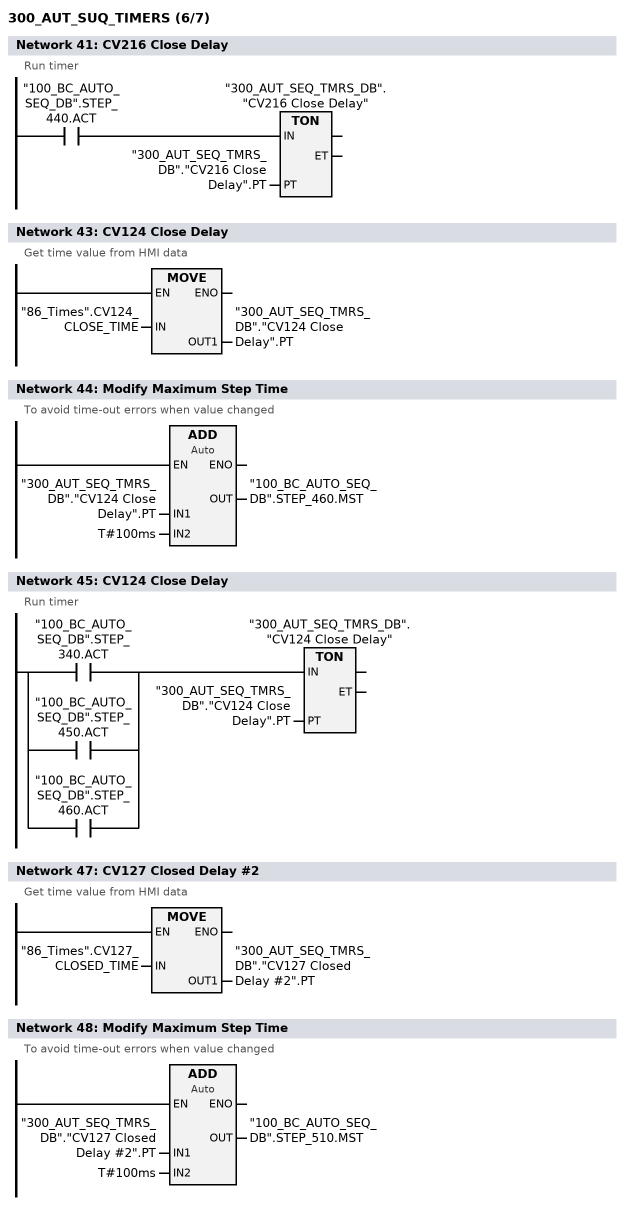
   "300_AUT_SEQ_TMRS_DB"."CV216 Close Delay".TON(IN := "100_BC_AUTO_SEQ_DB".STEP_440.ACT,
                           PT := "300_AUT_SEQ_TMRS_DB"."CV216 Close Delay".PT);
END_REGION

REGION Network 43: CV124 Close Delay
   // Get time value from HMI data
   RUNG wire#powerrail
      Move(in := "86_Times".CV124_CLOSE_TIME, out1 => "300_AUT_SEQ_TMRS_DB"."CV124 Close Delay".PT)
   END_RUNG
   // the same network as SCL:
   "300_AUT_SEQ_TMRS_DB"."CV124 Close Delay".PT := "86_Times".CV124_CLOSE_TIME;
END_REGION

REGION Network 44: Modify Maximum Step Time
   // To avoid time-out errors when value changed
   RUNG wire#powerrail
      Add(in1 := "300_AUT_SEQ_TMRS_DB"."CV124 Close Delay".PT, in2 := T#100ms, out => "100_BC_AUTO_SEQ_DB".STEP_460.MST)
   END_RUNG
   // the same network as SCL:
   "100_BC_AUTO_SEQ_DB".STEP_460.MST := "300_AUT_SEQ_TMRS_DB"."CV124 Close Delay".PT + T#100ms;
END_REGION

REGION Network 45: CV124 Close Delay
   // Run timer
   "300_AUT_SEQ_TMRS_DB"."CV124 Close Delay".TON(IN := "100_BC_AUTO_SEQ_DB".STEP_340.ACT OR "100_BC_AUTO_SEQ_DB".STEP_450.ACT OR "100_BC_AUTO_SEQ_DB".STEP_460.ACT,
                           PT := "300_AUT_SEQ_TMRS_DB"."CV124 Close Delay".PT);
END_REGION

REGION Network 47: CV127 Closed Delay #2
   // Get time value from HMI data
   RUNG wire#powerrail
      Move(in := "86_Times".CV127_CLOSED_TIME, out1 => "300_AUT_SEQ_TMRS_DB"."CV127 Closed Delay #2".PT)
   END_RUNG
   // the same network as SCL:
   "300_AUT_SEQ_TMRS_DB"."CV127 Closed Delay #2".PT := "86_Times".CV127_CLOSED_TIME;
END_REGION

REGION Network 48: Modify Maximum Step Time
   // To avoid time-out errors when value changed
   RUNG wire#powerrail
      Add(in1 := "300_AUT_SEQ_TMRS_DB"."CV127 Closed Delay #2".PT, in2 := T#100ms, out => "100_BC_AUTO_SEQ_DB".STEP_510.MST)
   END_RUNG
   // the same network as SCL:
   "100_BC_AUTO_SEQ_DB".STEP_510.MST := "300_AUT_SEQ_TMRS_DB"."CV127 Closed Delay #2".PT + T#100ms;
END_REGION

REGION Network 49: CV127 Closed Delay #2
   // Run timer
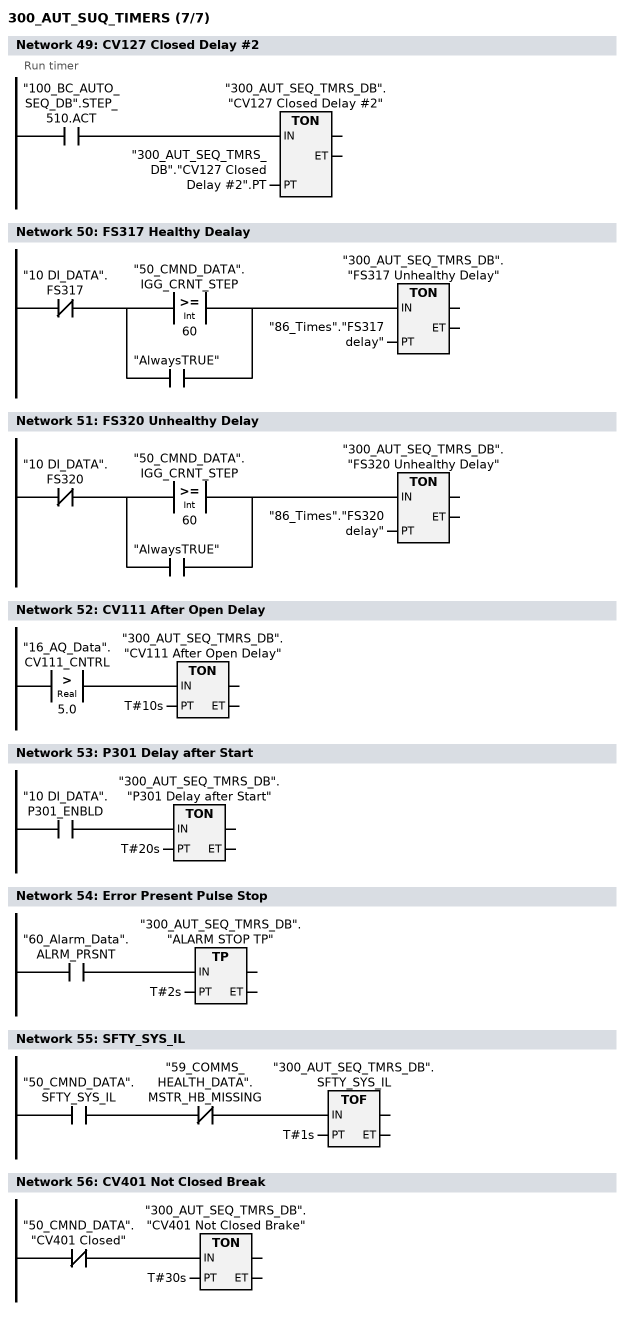
   "300_AUT_SEQ_TMRS_DB"."CV127 Closed Delay #2".TON(IN := "100_BC_AUTO_SEQ_DB".STEP_510.ACT,
                           PT := "300_AUT_SEQ_TMRS_DB"."CV127 Closed Delay #2".PT);
END_REGION

REGION Network 50: FS317 Healthy Dealay
   "300_AUT_SEQ_TMRS_DB"."FS317 Unhealthy Delay".TON(IN := NOT "10 DI_DATA".FS317 AND (("50_CMND_DATA".IGG_CRNT_STEP >= 60) OR "AlwaysTRUE"),
                           PT := "86_Times"."FS317 delay");
END_REGION

REGION Network 51: FS320 Unhealthy Delay
   "300_AUT_SEQ_TMRS_DB"."FS320 Unhealthy Delay".TON(IN := NOT "10 DI_DATA".FS320 AND (("50_CMND_DATA".IGG_CRNT_STEP >= 60) OR "AlwaysTRUE"),
                           PT := "86_Times"."FS320 delay");
END_REGION

REGION Network 52: CV111 After Open Delay
   "300_AUT_SEQ_TMRS_DB"."CV111 After Open Delay".TON(IN := "16_AQ_Data".CV111_CNTRL > 5.0, PT := T#10s);
END_REGION

REGION Network 53: P301 Delay after Start
   "300_AUT_SEQ_TMRS_DB"."P301 Delay after Start".TON(IN := "10 DI_DATA".P301_ENBLD, PT := T#20s);
END_REGION

REGION Network 54: Error Present Pulse Stop
   "300_AUT_SEQ_TMRS_DB"."ALARM STOP TP".TP(IN := "60_Alarm_Data".ALRM_PRSNT, PT := T#2s);
END_REGION

REGION Network 55: SFTY_SYS_IL
   "300_AUT_SEQ_TMRS_DB".SFTY_SYS_IL.TOF(IN := "50_CMND_DATA".SFTY_SYS_IL AND NOT "59_COMMS_HEALTH_DATA".MSTR_HB_MISSING,
                           PT := T#1s);
END_REGION

REGION Network 56: CV401 Not Closed Break
   "300_AUT_SEQ_TMRS_DB"."CV401 Not Closed Brake".TON(IN := NOT "50_CMND_DATA"."CV401 Closed", PT := T#30s);
END_REGION
END_FUNCTION

// folder: 50 - 59 PLC Communication

FUNCTION "51_GET_SLAVE_DATA" : Void   // FC51, LAD
TITLE = Get Slave Status Data
{ S7_Optimized_Access := 'TRUE' }
AUTHOR : JRS
VERSION : 0.1
// Code for getting status data from the slave PLC (IGG)
   VAR_TEMP
      RET_VAL_1 : Int;
   END_VAR
BEGIN

REGION Network 1: Get Slave Status Data
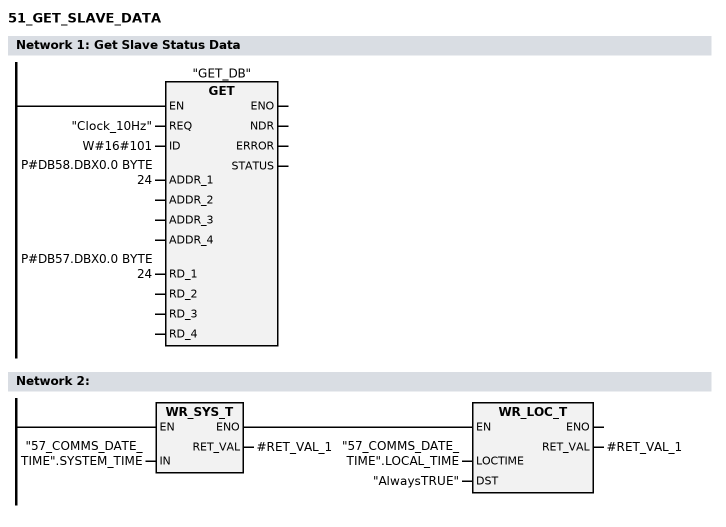
   "GET_DB"(REQ := "Clock_10Hz", ID := W#16#101, ADDR_1 := P#DB58.DBX0.0 BYTE 24, RD_1 := P#DB57.DBX0.0 BYTE 24);   // GET
END_REGION

REGION Network 2
   // ENO of a box is taken as its EN; it also drops when the box reports an error
   #RET_VAL_1 := WR_SYS_T(IN := "57_COMMS_DATE_TIME".SYSTEM_TIME);
   #RET_VAL_1 := WR_LOC_T(LOCTIME := "57_COMMS_DATE_TIME".LOCAL_TIME, DST := "AlwaysTRUE");
END_REGION
END_FUNCTION

FUNCTION "59_COMMS_HEALTH" : Void   // FC59, LAD
TITLE = Communications Heart Beats
{ S7_Optimized_Access := 'TRUE' }
AUTHOR : JRS
VERSION : 0.1
// Code for communications health determination
   VAR_TEMP   // added for the SCL form of the ladder/FBD networks
      _w1 : Bool;
   END_VAR
BEGIN

REGION Network 1: Local Heart Beat
   // Flip flop for status to other PLC's
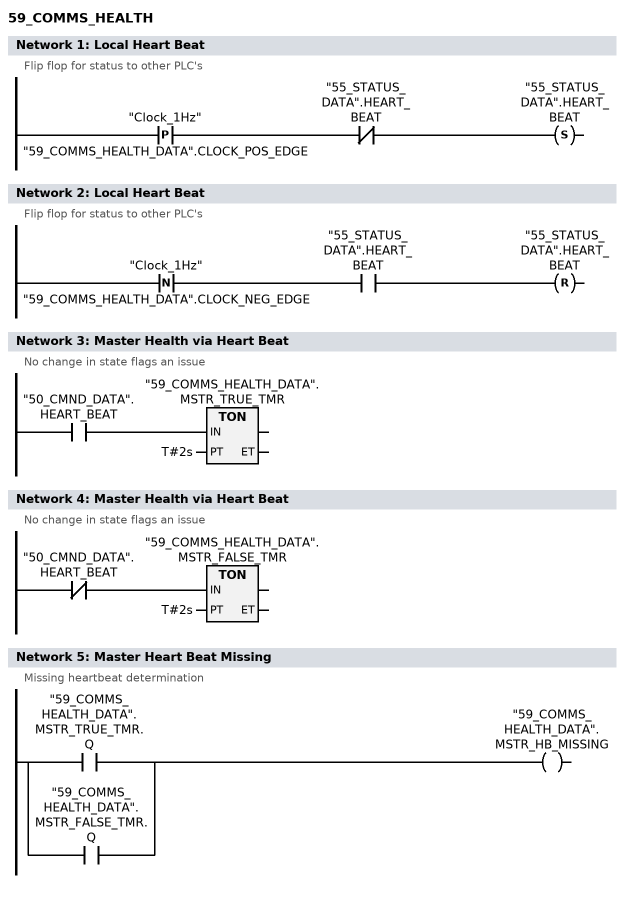
   RUNG wire#powerrail
      P_Contact(operand := "Clock_1Hz", bit := "59_COMMS_HEALTH_DATA".CLOCK_POS_EDGE)
      I_Contact( "55_STATUS_DATA".HEART_BEAT )
      S_Coil( "55_STATUS_DATA".HEART_BEAT )
   END_RUNG
   // the same network as SCL:
   #_w1 := "Clock_1Hz" AND NOT "59_COMMS_HEALTH_DATA".CLOCK_POS_EDGE;   // rising edge of "Clock_1Hz"
   "59_COMMS_HEALTH_DATA".CLOCK_POS_EDGE := "Clock_1Hz";
   IF #_w1 AND NOT "55_STATUS_DATA".HEART_BEAT THEN "55_STATUS_DATA".HEART_BEAT := TRUE; END_IF;
END_REGION

REGION Network 2: Local Heart Beat
   // Flip flop for status to other PLC's
   RUNG wire#powerrail
      N_Contact(operand := "Clock_1Hz", bit := "59_COMMS_HEALTH_DATA".CLOCK_NEG_EDGE)
      Contact( "55_STATUS_DATA".HEART_BEAT )
      R_Coil( "55_STATUS_DATA".HEART_BEAT )
   END_RUNG
   // the same network as SCL:
   #_w1 := NOT "Clock_1Hz" AND "59_COMMS_HEALTH_DATA".CLOCK_NEG_EDGE;   // falling edge of "Clock_1Hz"
   "59_COMMS_HEALTH_DATA".CLOCK_NEG_EDGE := "Clock_1Hz";
   IF #_w1 AND "55_STATUS_DATA".HEART_BEAT THEN "55_STATUS_DATA".HEART_BEAT := FALSE; END_IF;
END_REGION

REGION Network 3: Master Health via Heart Beat
   // No change in state flags an issue
   "59_COMMS_HEALTH_DATA".MSTR_TRUE_TMR.TON(IN := "50_CMND_DATA".HEART_BEAT, PT := T#2s);
END_REGION

REGION Network 4: Master Health via Heart Beat
   // No change in state flags an issue
   "59_COMMS_HEALTH_DATA".MSTR_FALSE_TMR.TON(IN := NOT "50_CMND_DATA".HEART_BEAT, PT := T#2s);
END_REGION

REGION Network 5: Master Heart Beat Missing
   // Missing heartbeat determination
   RUNG wire#powerrail
      Contact( "59_COMMS_HEALTH_DATA".MSTR_TRUE_TMR.Q )
      wire#w1
      Coil( "59_COMMS_HEALTH_DATA".MSTR_HB_MISSING )
   END_RUNG
   RUNG wire#powerrail
      Contact( "59_COMMS_HEALTH_DATA".MSTR_FALSE_TMR.Q )
   END_RUNG wire#w1
   // the same network as SCL:
   "59_COMMS_HEALTH_DATA".MSTR_HB_MISSING := "59_COMMS_HEALTH_DATA".MSTR_TRUE_TMR.Q OR "59_COMMS_HEALTH_DATA".MSTR_FALSE_TMR.Q;
END_REGION
END_FUNCTION

// folder: 500 - 699 Standard FBs

FUNCTION_BLOCK "500_SEQ_STEP"   // FB500, LAD
{ S7_Optimized_Access := 'TRUE' }
VERSION : 0.1
   VAR_INPUT
      SN : Int;   // Step number
      CS : Int;   // Current step
      MST : Time;   // Maximum step time
      SC : Bool;   // Step complete
      BPFLT : Bool;   // Bypass fault
   END_VAR
   VAR_OUTPUT
      ACT : Bool;   // Active
      DN : Bool;   // Done
   END_VAR
   VAR_IN_OUT
      AMST : Time;   // Actual maximum step time
      FLT : Bool;   // Timed out
   END_VAR
   VAR
      RNG : Bool;   // Running
   END_VAR
   VAR RETAIN
      STP_MAX_TIM : TON_TIME;   // Maximum step time
   END_VAR
BEGIN

REGION Network 1: Step Active
   // When step number is active, it is also running
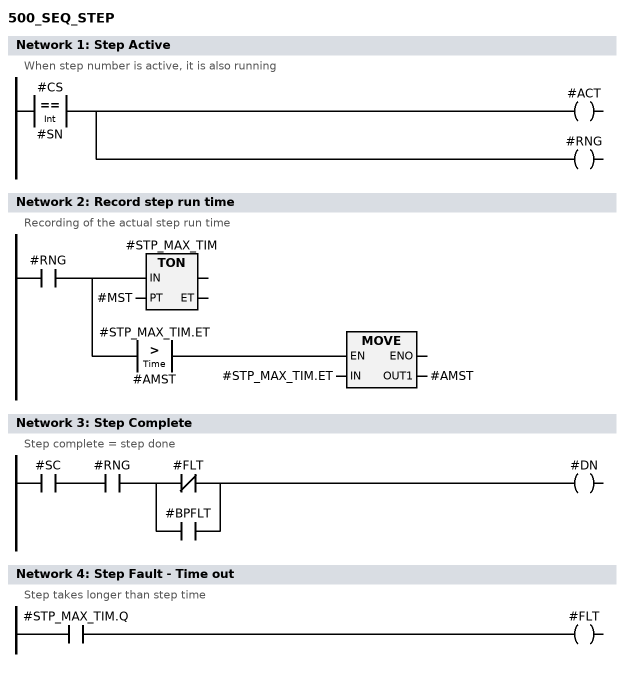
   RUNG wire#powerrail
      { S7_Templates := "SrcType := Int" } EQ_Contact(in1 := #CS, in2 := #SN)
      wire#w1
      Coil( #ACT )
   END_RUNG
   RUNG wire#w1
      Coil( #RNG )
   END_RUNG
   // the same network as SCL:
   #ACT := #CS = #SN;
   #RNG := #ACT;
END_REGION

REGION Network 2: Record step run time
   // Recording of the actual step run time
   #STP_MAX_TIM(IN := #RNG, PT := #MST);   // TON
   IF #RNG AND (#STP_MAX_TIM.ET > #AMST) THEN #AMST := #STP_MAX_TIM.ET; END_IF;
END_REGION

REGION Network 3: Step Complete
   // Step complete = step done
   RUNG wire#powerrail
      Contact( #SC )
      Contact( #RNG )
      wire#w1
      I_Contact( #FLT )
      wire#w2
      Coil( #DN )
   END_RUNG
   RUNG wire#w1
      Contact( #BPFLT )
   END_RUNG wire#w2
   // the same network as SCL:
   #DN := #SC AND #RNG AND (NOT #FLT OR #BPFLT);
END_REGION

REGION Network 4: Step Fault - Time out
   // Step takes longer than step time
   RUNG wire#powerrail
      Contact( #STP_MAX_TIM.Q )
      Coil( #FLT )
   END_RUNG
   // the same network as SCL:
   #FLT := #STP_MAX_TIM.Q;
END_REGION
END_FUNCTION_BLOCK

FUNCTION_BLOCK "64_Functioning Hours"   // FB501, LAD
{ S7_Optimized_Access := 'TRUE' }
VERSION : 0.1
   VAR_INPUT
      Started : Bool;
      Reset : Bool;
      "Service Time Days" : Int;
      "Service Time Hours" : Int;
   END_VAR
   VAR_OUTPUT
      Seconds : Int;
      Minutes : Int;
      Hours : Int;
      Days : Int;
      "Second beat_bit" : Bool;
      "Service Time bit" : Bool;
      "Hours to Service" : Int;
      "Hours Functioning Out" : Int;
      "Hours Total" : Int;
   END_VAR
   VAR
      "Second beat" : TON_TIME;
      "Second Reset" : TON_TIME;
   END_VAR
   VAR RETAIN
      "Seconds burn" : CTU_INT;
      "Minutes burn" : CTU_INT;
      "Hours burn" : CTU_INT;
      "Days burn" : CTU_INT;
      Aux : Struct
         Aux_1 : Bool;
         Aux_2 : Bool;
         Aux_3 : Bool;
         Aux_4 : Bool;
         Aux_Puls : Bool;
         Aux_PulsN : Bool;
         Aux_HoursFunctioning : Int;
         "Aux_Total Hours" : Int;
      END_STRUCT;
   END_VAR
   VAR
      "Hours Functioning" : Int;
   END_VAR
   VAR_TEMP   // added for the SCL form of the ladder/FBD networks
      _w1 : Bool;
      _w2 : Bool;
      _w3 : Bool;
   END_VAR
BEGIN

REGION Network 1
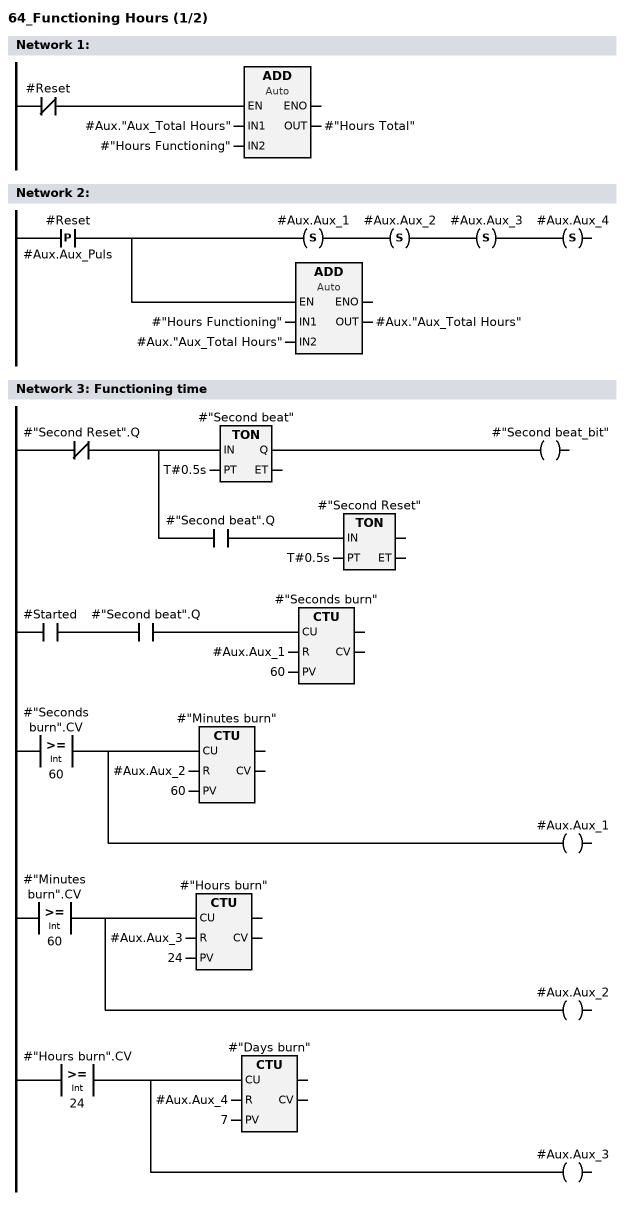
   RUNG wire#powerrail
      I_Contact( #Reset )
      Add(in1 := #Aux."Aux_Total Hours", in2 := #"Hours Functioning", out => #"Hours Total")
   END_RUNG
   // the same network as SCL:
   IF NOT #Reset THEN #"Hours Total" := #Aux."Aux_Total Hours" + #"Hours Functioning"; END_IF;
END_REGION

REGION Network 2
   RUNG wire#powerrail
      P_Contact(operand := #Reset, bit := #Aux.Aux_Puls)
      wire#w1
      S_Coil( #Aux.Aux_1 )
      S_Coil( #Aux.Aux_2 )
      S_Coil( #Aux.Aux_3 )
      S_Coil( #Aux.Aux_4 )
   END_RUNG
   RUNG wire#w1
      Add(in1 := #"Hours Functioning", in2 := #Aux."Aux_Total Hours", out => #Aux."Aux_Total Hours")
   END_RUNG
   // the same network as SCL:
   #_w1 := #Reset AND NOT #Aux.Aux_Puls;   // rising edge of #Reset
   #Aux.Aux_Puls := #Reset;
   IF #_w1 THEN
       #Aux.Aux_1 := TRUE;
       #Aux.Aux_2 := TRUE;
       #Aux.Aux_3 := TRUE;
       #Aux.Aux_4 := TRUE;
       #Aux."Aux_Total Hours" := #"Hours Functioning" + #Aux."Aux_Total Hours";
   END_IF;
END_REGION

REGION Network 3: Functioning time
   #"Second beat"(IN := NOT #"Second Reset".Q, PT := T#0.5s);   // TON
   #"Second beat_bit" := #"Second beat".Q;
   #"Second Reset"(IN := NOT #"Second Reset".Q AND #"Second beat".Q, PT := T#0.5s);   // TON
   #"Seconds burn"(CU := #Started AND #"Second beat".Q, R := #Aux.Aux_1, PV := 60);   // CTU
   #_w1 := #"Seconds burn".CV >= 60;
   #"Minutes burn"(CU := #_w1, R := #Aux.Aux_2, PV := 60);   // CTU
   #Aux.Aux_1 := #_w1;
   #_w2 := #"Minutes burn".CV >= 60;
   #"Hours burn"(CU := #_w2, R := #Aux.Aux_3, PV := 24);   // CTU
   #Aux.Aux_2 := #_w2;
   #_w3 := #"Hours burn".CV >= 24;
   #"Days burn"(CU := #_w3, R := #Aux.Aux_4, PV := 7);   // CTU
   #Aux.Aux_3 := #_w3;
END_REGION

REGION Network 4
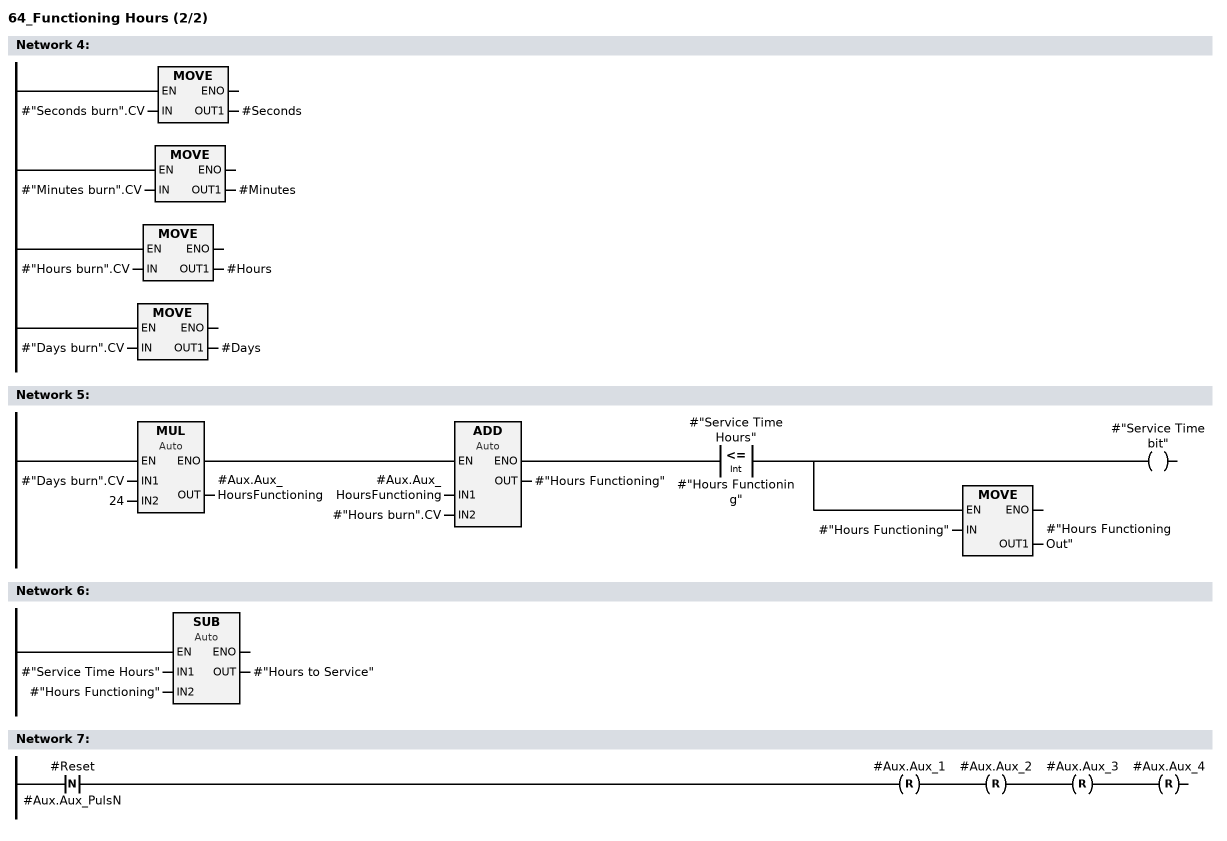
   RUNG wire#powerrail
      Move(in := #"Seconds burn".CV, out1 => #Seconds)
   END_RUNG
   RUNG wire#powerrail
      Move(in := #"Minutes burn".CV, out1 => #Minutes)
   END_RUNG
   RUNG wire#powerrail
      Move(in := #"Hours burn".CV, out1 => #Hours)
   END_RUNG
   RUNG wire#powerrail
      Move(in := #"Days burn".CV, out1 => #Days)
   END_RUNG
   // the same network as SCL:
   #Seconds := #"Seconds burn".CV;
   #Minutes := #"Minutes burn".CV;
   #Hours := #"Hours burn".CV;
   #Days := #"Days burn".CV;
END_REGION

REGION Network 5
   RUNG wire#powerrail
      Mul(in1 := #"Days burn".CV, in2 := 24, out => #Aux.Aux_HoursFunctioning)
      Add(in1 := #Aux.Aux_HoursFunctioning, in2 := #"Hours burn".CV, out => #"Hours Functioning")
      { S7_Templates := "SrcType := Int" } LE_Contact(in1 := #"Service Time Hours", in2 := #"Hours Functioning")
      wire#w1
      Coil( #"Service Time bit" )
   END_RUNG
   RUNG wire#w1
      Move(in := #"Hours Functioning", out1 => #"Hours Functioning Out")
   END_RUNG
   // the same network as SCL:
   #Aux.Aux_HoursFunctioning := #"Days burn".CV * 24;
   #"Hours Functioning" := #Aux.Aux_HoursFunctioning + #"Hours burn".CV;
   #"Service Time bit" := #"Service Time Hours" <= #"Hours Functioning";
   IF #"Service Time bit" THEN #"Hours Functioning Out" := #"Hours Functioning"; END_IF;
END_REGION

REGION Network 6
   RUNG wire#powerrail
      Sub(in1 := #"Service Time Hours", in2 := #"Hours Functioning", out => #"Hours to Service")
   END_RUNG
   // the same network as SCL:
   #"Hours to Service" := #"Service Time Hours" - #"Hours Functioning";
END_REGION

REGION Network 7
   RUNG wire#powerrail
      N_Contact(operand := #Reset, bit := #Aux.Aux_PulsN)
      R_Coil( #Aux.Aux_1 )
      R_Coil( #Aux.Aux_2 )
      R_Coil( #Aux.Aux_3 )
      R_Coil( #Aux.Aux_4 )
   END_RUNG
   // the same network as SCL:
   #_w1 := NOT #Reset AND #Aux.Aux_PulsN;   // falling edge of #Reset
   #Aux.Aux_PulsN := #Reset;
   IF #_w1 THEN
       #Aux.Aux_1 := FALSE;
       #Aux.Aux_2 := FALSE;
       #Aux.Aux_3 := FALSE;
       #Aux.Aux_4 := FALSE;
   END_IF;
END_REGION
END_FUNCTION_BLOCK

FUNCTION_BLOCK "502_ALM_ANALOG"   // FB502, LAD
{ S7_Optimized_Access := 'FALSE' }